REGION Network 19: TURUNKAN PRESSURE V 5
   RUNG wire#powerrail
      Contact( "DB106".Out_Step_17 )
      wire#w1
      I_Contact( "DB106".En_Step_19 )
      I_Contact( "Emergency" )
      Coil( "DB106".En_Step_18 )
   END_RUNG
   RUNG wire#powerrail
      Contact( "DB106".En_Step_18 )
   END_RUNG wire#w1
   // the same network as SCL:
   "DB106".En_Step_18 := ("DB106".Out_Step_17 OR "DB106".En_Step_18) AND NOT "DB106".En_Step_19 AND NOT "Emergency";
END_REGION

REGION Network 20: VB 5 OFF
   RUNG wire#powerrail
      Contact( "DB106".Out_Step_18 )
      { S7_Templates := "SrcType := Int" } LT_Contact(in1 := "Pressure vessel 5", in2 := 3)
      wire#w1
      I_Contact( "DB106".En_Step_20 )
      I_Contact( "Emergency" )
      Coil( "DB106".En_Step_19 )
   END_RUNG
   RUNG wire#powerrail
      Contact( "DB106".En_Step_19 )
   END_RUNG wire#w1
   // the same network as SCL:
   "DB106".En_Step_19 := (("DB106".Out_Step_18 AND ("Pressure vessel 5" < 3)) OR "DB106".En_Step_19) AND NOT "DB106".En_Step_20 AND NOT "Emergency";
END_REGION

REGION Network 21: VP 86 ON VP OFF
   RUNG wire#powerrail
      Contact( "DB106".Out_Step_19 )
      S_ODT(T_NO := "Tag_88", TV := S5T#4S, R :=, BI =>, RET_VAL =>)
      wire#w1
      I_Contact( "DB106".En_Step_21 )
      I_Contact( "Emergency" )
      Coil( "DB106".En_Step_20 )
   END_RUNG
   RUNG wire#powerrail
      Contact( "DB106".En_Step_20 )
   END_RUNG wire#w1
   // the same network as SCL:
   #_s5time1 := S_ODT(T_NO := "Tag_88", S := "DB106".Out_Step_19, TV := S5T#4S, Q => #_w1);
   "DB106".En_Step_20 := (#_w1 OR "DB106".En_Step_20) AND NOT "DB106".En_Step_21 AND NOT "Emergency";
END_REGION

REGION Network 22: VP 86 OFF VP 87 ON
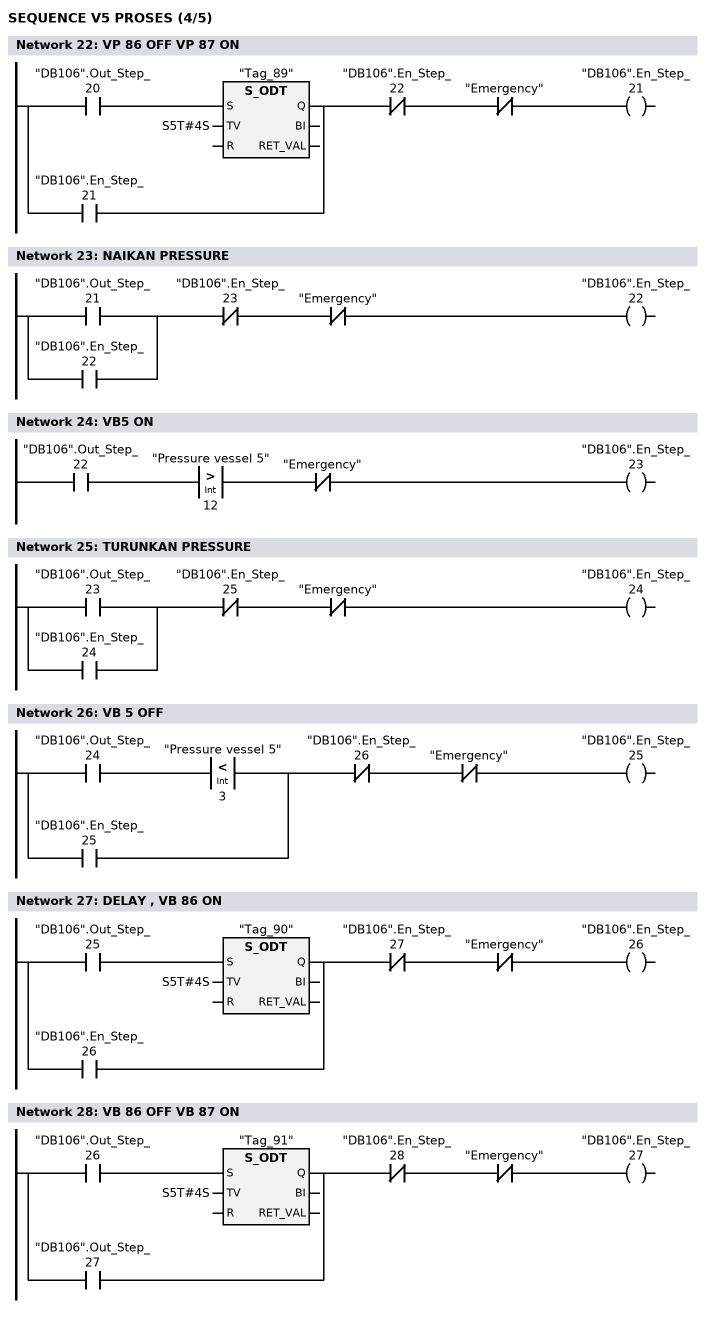
   RUNG wire#powerrail
      Contact( "DB106".Out_Step_20 )
      S_ODT(T_NO := "Tag_89", TV := S5T#4S, R :=, BI =>, RET_VAL =>)
      wire#w1
      I_Contact( "DB106".En_Step_22 )
      I_Contact( "Emergency" )
      Coil( "DB106".En_Step_21 )
   END_RUNG
   RUNG wire#powerrail
      Contact( "DB106".En_Step_21 )
   END_RUNG wire#w1
   // the same network as SCL:
   #_s5time1 := S_ODT(T_NO := "Tag_89", S := "DB106".Out_Step_20, TV := S5T#4S, Q => #_w1);
   "DB106".En_Step_21 := (#_w1 OR "DB106".En_Step_21) AND NOT "DB106".En_Step_22 AND NOT "Emergency";
END_REGION

REGION Network 23: NAIKAN PRESSURE
   RUNG wire#powerrail
      Contact( "DB106".Out_Step_21 )
      wire#w1
      I_Contact( "DB106".En_Step_23 )
      I_Contact( "Emergency" )
      Coil( "DB106".En_Step_22 )
   END_RUNG
   RUNG wire#powerrail
      Contact( "DB106".En_Step_22 )
   END_RUNG wire#w1
   // the same network as SCL:
   "DB106".En_Step_22 := ("DB106".Out_Step_21 OR "DB106".En_Step_22) AND NOT "DB106".En_Step_23 AND NOT "Emergency";
END_REGION

REGION Network 24: VB5 ON
   RUNG wire#powerrail
      Contact( "DB106".Out_Step_22 )
      { S7_Templates := "SrcType := Int" } GT_Contact(in1 := "Pressure vessel 5", in2 := 12)
      I_Contact( "Emergency" )
      Coil( "DB106".En_Step_23 )
   END_RUNG
   // the same network as SCL:
   "DB106".En_Step_23 := "DB106".Out_Step_22 AND ("Pressure vessel 5" > 12) AND NOT "Emergency";
END_REGION

REGION Network 25: TURUNKAN PRESSURE
   RUNG wire#powerrail
      Contact( "DB106".Out_Step_23 )
      wire#w1
      I_Contact( "DB106".En_Step_25 )
      I_Contact( "Emergency" )
      Coil( "DB106".En_Step_24 )
   END_RUNG
   RUNG wire#powerrail
      Contact( "DB106".En_Step_24 )
   END_RUNG wire#w1
   // the same network as SCL:
   "DB106".En_Step_24 := ("DB106".Out_Step_23 OR "DB106".En_Step_24) AND NOT "DB106".En_Step_25 AND NOT "Emergency";
END_REGION

REGION Network 26: VB 5 OFF
   RUNG wire#powerrail
      Contact( "DB106".Out_Step_24 )
      { S7_Templates := "SrcType := Int" } LT_Contact(in1 := "Pressure vessel 5", in2 := 3)
      wire#w1
      I_Contact( "DB106".En_Step_26 )
      I_Contact( "Emergency" )
      Coil( "DB106".En_Step_25 )
   END_RUNG
   RUNG wire#powerrail
      Contact( "DB106".En_Step_25 )
   END_RUNG wire#w1
   // the same network as SCL:
   "DB106".En_Step_25 := (("DB106".Out_Step_24 AND ("Pressure vessel 5" < 3)) OR "DB106".En_Step_25) AND NOT "DB106".En_Step_26 AND NOT "Emergency";
END_REGION

REGION Network 27: DELAY , VB 86 ON
   RUNG wire#powerrail
      Contact( "DB106".Out_Step_25 )
      S_ODT(T_NO := "Tag_90", TV := S5T#4S, R :=, BI =>, RET_VAL =>)
      wire#w1
      I_Contact( "DB106".En_Step_27 )
      I_Contact( "Emergency" )
      Coil( "DB106".En_Step_26 )
   END_RUNG
   RUNG wire#powerrail
      Contact( "DB106".En_Step_26 )
   END_RUNG wire#w1
   // the same network as SCL:
   #_s5time1 := S_ODT(T_NO := "Tag_90", S := "DB106".Out_Step_25, TV := S5T#4S, Q => #_w1);
   "DB106".En_Step_26 := (#_w1 OR "DB106".En_Step_26) AND NOT "DB106".En_Step_27 AND NOT "Emergency";
END_REGION

REGION Network 28: VB 86 OFF VB 87 ON
   RUNG wire#powerrail
      Contact( "DB106".Out_Step_26 )
      S_ODT(T_NO := "Tag_91", TV := S5T#4S, R :=, BI =>, RET_VAL =>)
      wire#w1
      I_Contact( "DB106".En_Step_28 )
      I_Contact( "Emergency" )
      Coil( "DB106".En_Step_27 )
   END_RUNG
   RUNG wire#powerrail
      Contact( "DB106".Out_Step_27 )
   END_RUNG wire#w1
   // the same network as SCL:
   #_s5time1 := S_ODT(T_NO := "Tag_91", S := "DB106".Out_Step_26, TV := S5T#4S, Q => #_w1);
   "DB106".En_Step_27 := (#_w1 OR "DB106".Out_Step_27) AND NOT "DB106".En_Step_28 AND NOT "Emergency";
END_REGION

REGION Network 29
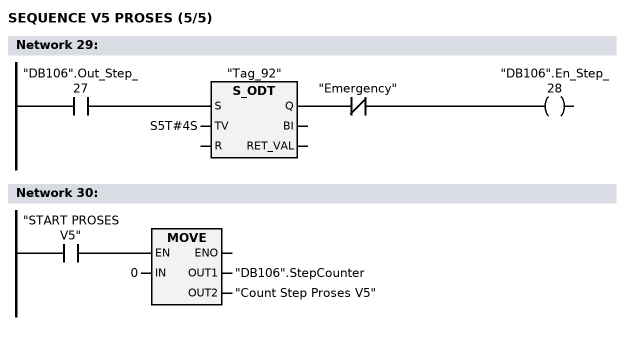
   RUNG wire#powerrail
      Contact( "DB106".Out_Step_27 )
      S_ODT(T_NO := "Tag_92", TV := S5T#4S, R :=, BI =>, RET_VAL =>)
      I_Contact( "Emergency" )
      Coil( "DB106".En_Step_28 )
   END_RUNG
   // the same network as SCL:
   #_s5time1 := S_ODT(T_NO := "Tag_92", S := "DB106".Out_Step_27, TV := S5T#4S, Q => #_w1);
   "DB106".En_Step_28 := #_w1 AND NOT "Emergency";
END_REGION

REGION Network 30
   RUNG wire#powerrail
      Contact( "START PROSES V5" )
      Move(in := 0, out1 => "DB106".StepCounter, out2 => "Count Step Proses V5")
   END_RUNG
   // the same network as SCL:
   IF "START PROSES V5" THEN
       "DB106".StepCounter := 0;
       "Count Step Proses V5" := 0;
   END_IF;
END_REGION
END_FUNCTION

FUNCTION "VESSEL 6 PROSES" : Void   // FC19, LAD
{ S7_Optimized_Access := 'TRUE' }
VERSION : 0.1
   VAR_TEMP   // added for the SCL form of the ladder/FBD networks
      _w1 : Bool;
      _w2 : Bool;
   END_VAR
BEGIN

REGION Network 1
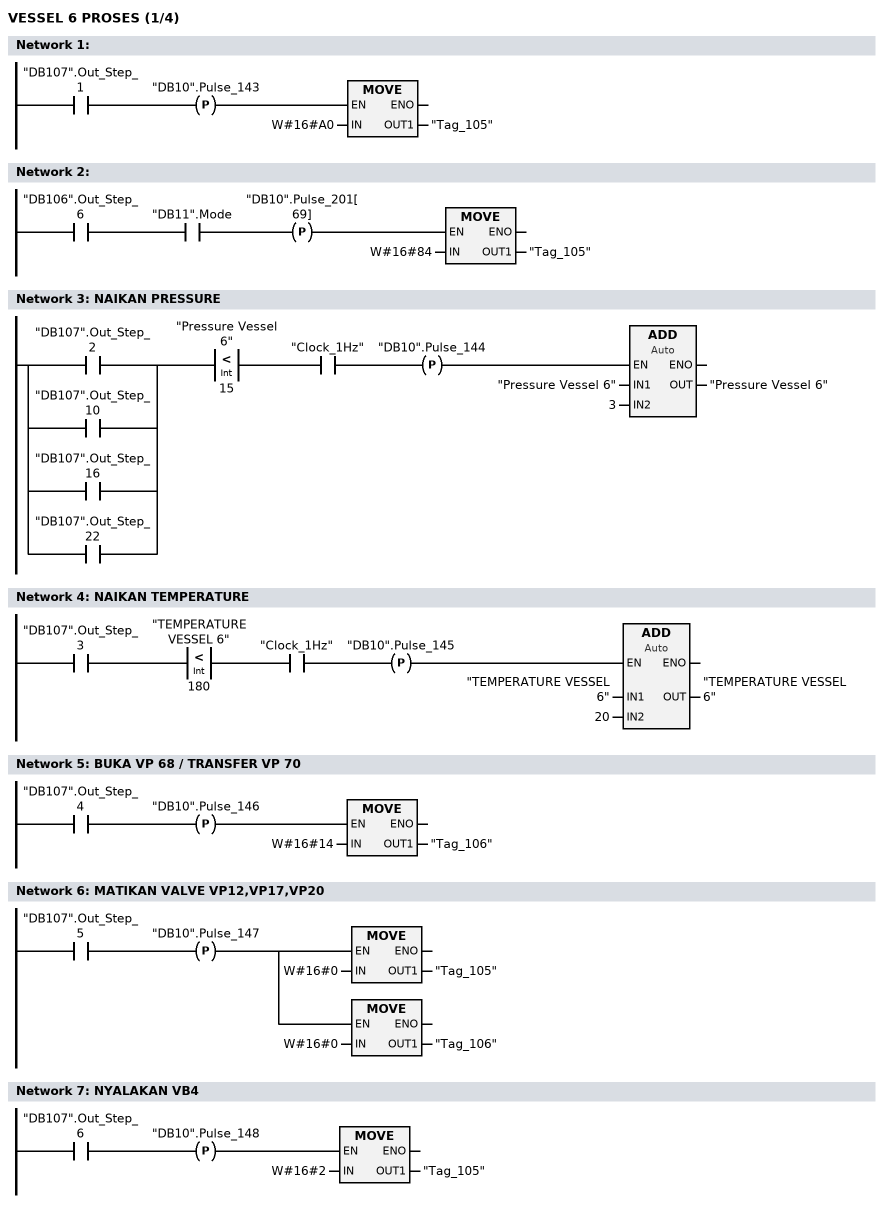
   RUNG wire#powerrail
      Contact( "DB107".Out_Step_1 )
      P_Trig( "DB10".Pulse_143 )
      Move(in := W#16#A0, out1 => "Tag_105")
   END_RUNG
   // the same network as SCL:
   #_w1 := "DB107".Out_Step_1 AND NOT "DB10".Pulse_143;   // rising edge
   "DB10".Pulse_143 := "DB107".Out_Step_1;
   IF #_w1 THEN "Tag_105" := W#16#A0; END_IF;
END_REGION

REGION Network 2
   RUNG wire#powerrail
      Contact( "DB106".Out_Step_6 )
      Contact( "DB11".Mode )
      P_Trig( "DB10".Pulse_201[69] )
      Move(in := W#16#84, out1 => "Tag_105")
   END_RUNG
   // the same network as SCL:
   #_w1 := "DB106".Out_Step_6 AND "DB11".Mode;
   #_w2 := #_w1 AND NOT "DB10".Pulse_201[69];   // rising edge
   "DB10".Pulse_201[69] := #_w1;
   IF #_w2 THEN "Tag_105" := W#16#84; END_IF;
END_REGION

REGION Network 3: NAIKAN PRESSURE
   RUNG wire#powerrail
      Contact( "DB107".Out_Step_2 )
      wire#w1
      { S7_Templates := "SrcType := Int" } LT_Contact(in1 := "Pressure Vessel 6", in2 := 15)
      Contact( "Clock_1Hz" )
      P_Trig( "DB10".Pulse_144 )
      Add(in1 := "Pressure Vessel 6", in2 := 3, out => "Pressure Vessel 6")
   END_RUNG
   RUNG wire#powerrail
      Contact( "DB107".Out_Step_10 )
   END_RUNG wire#w1
   RUNG wire#powerrail
      Contact( "DB107".Out_Step_16 )
   END_RUNG wire#w1
   RUNG wire#powerrail
      Contact( "DB107".Out_Step_22 )
   END_RUNG wire#w1
   // the same network as SCL:
   #_w1 := ("DB107".Out_Step_2 OR "DB107".Out_Step_10 OR "DB107".Out_Step_16 OR "DB107".Out_Step_22) AND ("Pressure Vessel 6" < 15) AND "Clock_1Hz";
   #_w2 := #_w1 AND NOT "DB10".Pulse_144;   // rising edge
   "DB10".Pulse_144 := #_w1;
   IF #_w2 THEN "Pressure Vessel 6" := "Pressure Vessel 6" + 3; END_IF;
END_REGION

REGION Network 4: NAIKAN TEMPERATURE
   RUNG wire#powerrail
      Contact( "DB107".Out_Step_3 )
      { S7_Templates := "SrcType := Int" } LT_Contact(in1 := "TEMPERATURE VESSEL 6", in2 := 180)
      Contact( "Clock_1Hz" )
      P_Trig( "DB10".Pulse_145 )
      Add(in1 := "TEMPERATURE VESSEL 6", in2 := 20, out => "TEMPERATURE VESSEL 6")
   END_RUNG
   // the same network as SCL:
   #_w1 := "DB107".Out_Step_3 AND ("TEMPERATURE VESSEL 6" < 180) AND "Clock_1Hz";
   #_w2 := #_w1 AND NOT "DB10".Pulse_145;   // rising edge
   "DB10".Pulse_145 := #_w1;
   IF #_w2 THEN "TEMPERATURE VESSEL 6" := "TEMPERATURE VESSEL 6" + 20; END_IF;
END_REGION

REGION Network 5: BUKA VP 68 / TRANSFER VP 70
   RUNG wire#powerrail
      Contact( "DB107".Out_Step_4 )
      P_Trig( "DB10".Pulse_146 )
      Move(in := W#16#14, out1 => "Tag_106")
   END_RUNG
   // the same network as SCL:
   #_w1 := "DB107".Out_Step_4 AND NOT "DB10".Pulse_146;   // rising edge
   "DB10".Pulse_146 := "DB107".Out_Step_4;
   IF #_w1 THEN "Tag_106" := W#16#14; END_IF;
END_REGION

REGION Network 6: MATIKAN VALVE VP12,VP17,VP20
   RUNG wire#powerrail
      Contact( "DB107".Out_Step_5 )
      P_Trig( "DB10".Pulse_147 )
      wire#w1
      Move(in := W#16#0, out1 => "Tag_105")
   END_RUNG
   RUNG wire#w1
      Move(in := W#16#0, out1 => "Tag_106")
   END_RUNG
   // the same network as SCL:
   #_w1 := "DB107".Out_Step_5 AND NOT "DB10".Pulse_147;   // rising edge
   "DB10".Pulse_147 := "DB107".Out_Step_5;
   IF #_w1 THEN
       "Tag_105" := W#16#0;
       "Tag_106" := W#16#0;
   END_IF;
END_REGION

REGION Network 7: NYALAKAN VB4
   RUNG wire#powerrail
      Contact( "DB107".Out_Step_6 )
      P_Trig( "DB10".Pulse_148 )
      Move(in := W#16#2, out1 => "Tag_105")
   END_RUNG
   // the same network as SCL:
   #_w1 := "DB107".Out_Step_6 AND NOT "DB10".Pulse_148;   // rising edge
   "DB10".Pulse_148 := "DB107".Out_Step_6;
   IF #_w1 THEN "Tag_105" := W#16#2; END_IF;
END_REGION

REGION Network 8: TURUNKAN PRESSURE
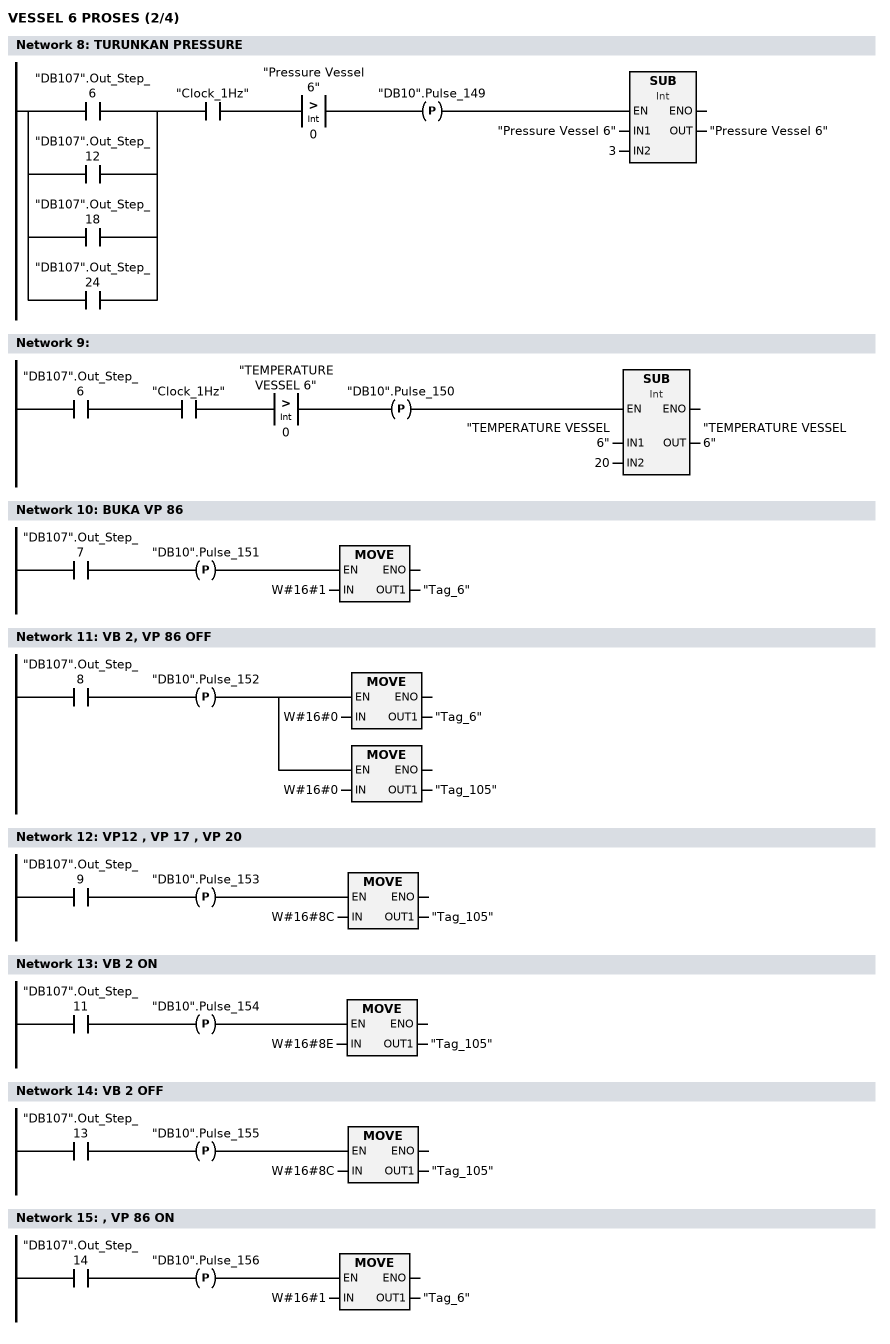
   RUNG wire#powerrail
      Contact( "DB107".Out_Step_6 )
      wire#w1
      Contact( "Clock_1Hz" )
      { S7_Templates := "SrcType := Int" } GT_Contact(in1 := "Pressure Vessel 6", in2 := 0)
      P_Trig( "DB10".Pulse_149 )
      { S7_Templates := "SrcType := Int" } Sub(in1 := "Pressure Vessel 6", in2 := 3, out => "Pressure Vessel 6")
   END_RUNG
   RUNG wire#powerrail
      Contact( "DB107".Out_Step_12 )
   END_RUNG wire#w1
   RUNG wire#powerrail
      Contact( "DB107".Out_Step_18 )
   END_RUNG wire#w1
   RUNG wire#powerrail
      Contact( "DB107".Out_Step_24 )
   END_RUNG wire#w1
   // the same network as SCL:
   #_w1 := ("DB107".Out_Step_6 OR "DB107".Out_Step_12 OR "DB107".Out_Step_18 OR "DB107".Out_Step_24) AND "Clock_1Hz" AND ("Pressure Vessel 6" > 0);
   #_w2 := #_w1 AND NOT "DB10".Pulse_149;   // rising edge
   "DB10".Pulse_149 := #_w1;
   IF #_w2 THEN "Pressure Vessel 6" := "Pressure Vessel 6" - 3; END_IF;
END_REGION

REGION Network 9
   RUNG wire#powerrail
      Contact( "DB107".Out_Step_6 )
      Contact( "Clock_1Hz" )
      { S7_Templates := "SrcType := Int" } GT_Contact(in1 := "TEMPERATURE VESSEL 6", in2 := 0)
      P_Trig( "DB10".Pulse_150 )
      { S7_Templates := "SrcType := Int" } Sub(in1 := "TEMPERATURE VESSEL 6", in2 := 20, out => "TEMPERATURE VESSEL 6")
   END_RUNG
   // the same network as SCL:
   #_w1 := "DB107".Out_Step_6 AND "Clock_1Hz" AND ("TEMPERATURE VESSEL 6" > 0);
   #_w2 := #_w1 AND NOT "DB10".Pulse_150;   // rising edge
   "DB10".Pulse_150 := #_w1;
   IF #_w2 THEN "TEMPERATURE VESSEL 6" := "TEMPERATURE VESSEL 6" - 20; END_IF;
END_REGION

REGION Network 10: BUKA VP 86
   RUNG wire#powerrail
      Contact( "DB107".Out_Step_7 )
      P_Trig( "DB10".Pulse_151 )
      Move(in := W#16#1, out1 => "Tag_6")
   END_RUNG
   // the same network as SCL:
   #_w1 := "DB107".Out_Step_7 AND NOT "DB10".Pulse_151;   // rising edge
   "DB10".Pulse_151 := "DB107".Out_Step_7;
   IF #_w1 THEN "Tag_6" := W#16#1; END_IF;
END_REGION

REGION Network 11: VB 2, VP 86 OFF
   RUNG wire#powerrail
      Contact( "DB107".Out_Step_8 )
      P_Trig( "DB10".Pulse_152 )
      wire#w1
      Move(in := W#16#0, out1 => "Tag_6")
   END_RUNG
   RUNG wire#w1
      Move(in := W#16#0, out1 => "Tag_105")
   END_RUNG
   // the same network as SCL:
   #_w1 := "DB107".Out_Step_8 AND NOT "DB10".Pulse_152;   // rising edge
   "DB10".Pulse_152 := "DB107".Out_Step_8;
   IF #_w1 THEN
       "Tag_6" := W#16#0;
       "Tag_105" := W#16#0;
   END_IF;
END_REGION

REGION Network 12: VP12 , VP 17 , VP 20
   RUNG wire#powerrail
      Contact( "DB107".Out_Step_9 )
      P_Trig( "DB10".Pulse_153 )
      Move(in := W#16#8C, out1 => "Tag_105")
   END_RUNG
   // the same network as SCL:
   #_w1 := "DB107".Out_Step_9 AND NOT "DB10".Pulse_153;   // rising edge
   "DB10".Pulse_153 := "DB107".Out_Step_9;
   IF #_w1 THEN "Tag_105" := W#16#8C; END_IF;
END_REGION

REGION Network 13: VB 2 ON
   RUNG wire#powerrail
      Contact( "DB107".Out_Step_11 )
      P_Trig( "DB10".Pulse_154 )
      Move(in := W#16#8E, out1 => "Tag_105")
   END_RUNG
   // the same network as SCL:
   #_w1 := "DB107".Out_Step_11 AND NOT "DB10".Pulse_154;   // rising edge
   "DB10".Pulse_154 := "DB107".Out_Step_11;
   IF #_w1 THEN "Tag_105" := W#16#8E; END_IF;
END_REGION

REGION Network 14: VB 2 OFF
   RUNG wire#powerrail
      Contact( "DB107".Out_Step_13 )
      P_Trig( "DB10".Pulse_155 )
      Move(in := W#16#8C, out1 => "Tag_105")
   END_RUNG
   // the same network as SCL:
   #_w1 := "DB107".Out_Step_13 AND NOT "DB10".Pulse_155;   // rising edge
   "DB10".Pulse_155 := "DB107".Out_Step_13;
   IF #_w1 THEN "Tag_105" := W#16#8C; END_IF;
END_REGION

REGION Network 15: , VP 86 ON
   RUNG wire#powerrail
      Contact( "DB107".Out_Step_14 )
      P_Trig( "DB10".Pulse_156 )
      Move(in := W#16#1, out1 => "Tag_6")
   END_RUNG
   // the same network as SCL:
   #_w1 := "DB107".Out_Step_14 AND NOT "DB10".Pulse_156;   // rising edge
   "DB10".Pulse_156 := "DB107".Out_Step_14;
   IF #_w1 THEN "Tag_6" := W#16#1; END_IF;
END_REGION

REGION Network 16: VP 86 OFF
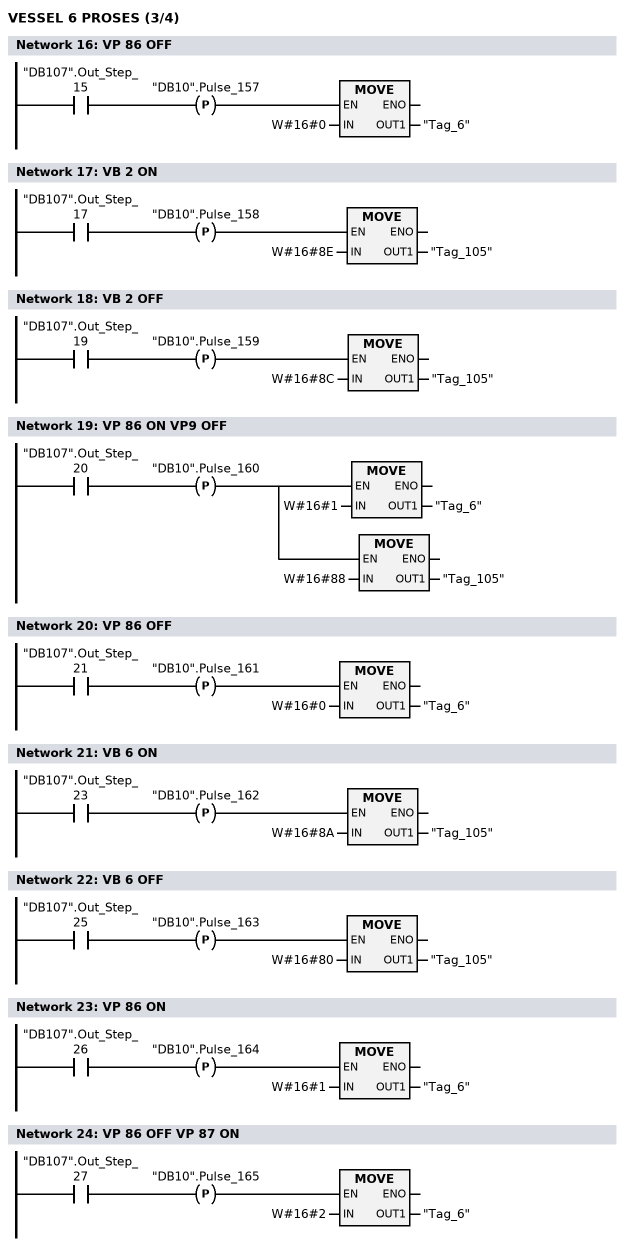
   RUNG wire#powerrail
      Contact( "DB107".Out_Step_15 )
      P_Trig( "DB10".Pulse_157 )
      Move(in := W#16#0, out1 => "Tag_6")
   END_RUNG
   // the same network as SCL:
   #_w1 := "DB107".Out_Step_15 AND NOT "DB10".Pulse_157;   // rising edge
   "DB10".Pulse_157 := "DB107".Out_Step_15;
   IF #_w1 THEN "Tag_6" := W#16#0; END_IF;
END_REGION

REGION Network 17: VB 2 ON
   RUNG wire#powerrail
      Contact( "DB107".Out_Step_17 )
      P_Trig( "DB10".Pulse_158 )
      Move(in := W#16#8E, out1 => "Tag_105")
   END_RUNG
   // the same network as SCL:
   #_w1 := "DB107".Out_Step_17 AND NOT "DB10".Pulse_158;   // rising edge
   "DB10".Pulse_158 := "DB107".Out_Step_17;
   IF #_w1 THEN "Tag_105" := W#16#8E; END_IF;
END_REGION

REGION Network 18: VB 2 OFF
   RUNG wire#powerrail
      Contact( "DB107".Out_Step_19 )
      P_Trig( "DB10".Pulse_159 )
      Move(in := W#16#8C, out1 => "Tag_105")
   END_RUNG
   // the same network as SCL:
   #_w1 := "DB107".Out_Step_19 AND NOT "DB10".Pulse_159;   // rising edge
   "DB10".Pulse_159 := "DB107".Out_Step_19;
   IF #_w1 THEN "Tag_105" := W#16#8C; END_IF;
END_REGION

REGION Network 19: VP 86 ON VP9 OFF
   RUNG wire#powerrail
      Contact( "DB107".Out_Step_20 )
      P_Trig( "DB10".Pulse_160 )
      wire#w1
      Move(in := W#16#1, out1 => "Tag_6")
   END_RUNG
   RUNG wire#w1
      Move(in := W#16#88, out1 => "Tag_105")
   END_RUNG
   // the same network as SCL:
   #_w1 := "DB107".Out_Step_20 AND NOT "DB10".Pulse_160;   // rising edge
   "DB10".Pulse_160 := "DB107".Out_Step_20;
   IF #_w1 THEN
       "Tag_6" := W#16#1;
       "Tag_105" := W#16#88;
   END_IF;
END_REGION

REGION Network 20: VP 86 OFF
   RUNG wire#powerrail
      Contact( "DB107".Out_Step_21 )
      P_Trig( "DB10".Pulse_161 )
      Move(in := W#16#0, out1 => "Tag_6")
   END_RUNG
   // the same network as SCL:
   #_w1 := "DB107".Out_Step_21 AND NOT "DB10".Pulse_161;   // rising edge
   "DB10".Pulse_161 := "DB107".Out_Step_21;
   IF #_w1 THEN "Tag_6" := W#16#0; END_IF;
END_REGION

REGION Network 21: VB 6 ON
   RUNG wire#powerrail
      Contact( "DB107".Out_Step_23 )
      P_Trig( "DB10".Pulse_162 )
      Move(in := W#16#8A, out1 => "Tag_105")
   END_RUNG
   // the same network as SCL:
   #_w1 := "DB107".Out_Step_23 AND NOT "DB10".Pulse_162;   // rising edge
   "DB10".Pulse_162 := "DB107".Out_Step_23;
   IF #_w1 THEN "Tag_105" := W#16#8A; END_IF;
END_REGION

REGION Network 22: VB 6 OFF
   RUNG wire#powerrail
      Contact( "DB107".Out_Step_25 )
      P_Trig( "DB10".Pulse_163 )
      Move(in := W#16#80, out1 => "Tag_105")
   END_RUNG
   // the same network as SCL:
   #_w1 := "DB107".Out_Step_25 AND NOT "DB10".Pulse_163;   // rising edge
   "DB10".Pulse_163 := "DB107".Out_Step_25;
   IF #_w1 THEN "Tag_105" := W#16#80; END_IF;
END_REGION

REGION Network 23: VP 86 ON
   RUNG wire#powerrail
      Contact( "DB107".Out_Step_26 )
      P_Trig( "DB10".Pulse_164 )
      Move(in := W#16#1, out1 => "Tag_6")
   END_RUNG
   // the same network as SCL:
   #_w1 := "DB107".Out_Step_26 AND NOT "DB10".Pulse_164;   // rising edge
   "DB10".Pulse_164 := "DB107".Out_Step_26;
   IF #_w1 THEN "Tag_6" := W#16#1; END_IF;
END_REGION

REGION Network 24: VP 86 OFF VP 87 ON
   RUNG wire#powerrail
      Contact( "DB107".Out_Step_27 )
      P_Trig( "DB10".Pulse_165 )
      Move(in := W#16#2, out1 => "Tag_6")
   END_RUNG
   // the same network as SCL:
   #_w1 := "DB107".Out_Step_27 AND NOT "DB10".Pulse_165;   // rising edge
   "DB10".Pulse_165 := "DB107".Out_Step_27;
   IF #_w1 THEN "Tag_6" := W#16#2; END_IF;
END_REGION

REGION Network 25: VP 87 OFF
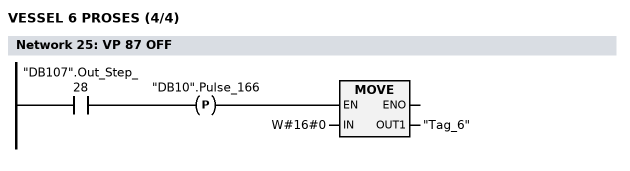
   RUNG wire#powerrail
      Contact( "DB107".Out_Step_28 )
      P_Trig( "DB10".Pulse_166 )
      Move(in := W#16#0, out1 => "Tag_6")
   END_RUNG
   // the same network as SCL:
   #_w1 := "DB107".Out_Step_28 AND NOT "DB10".Pulse_166;   // rising edge
   "DB10".Pulse_166 := "DB107".Out_Step_28;
   IF #_w1 THEN "Tag_6" := W#16#0; END_IF;
END_REGION
END_FUNCTION

FUNCTION "SEQUENCE V6 PROSES" : Void   // FC20, LAD
{ S7_Optimized_Access := 'TRUE' }
VERSION : 0.1
   VAR_TEMP   // added for the SCL form of the ladder/FBD networks
      _w1 : Bool;
      _w2 : Bool;
      _s5time1 : S5Time;
   END_VAR
BEGIN

REGION Network 1: START PROSES
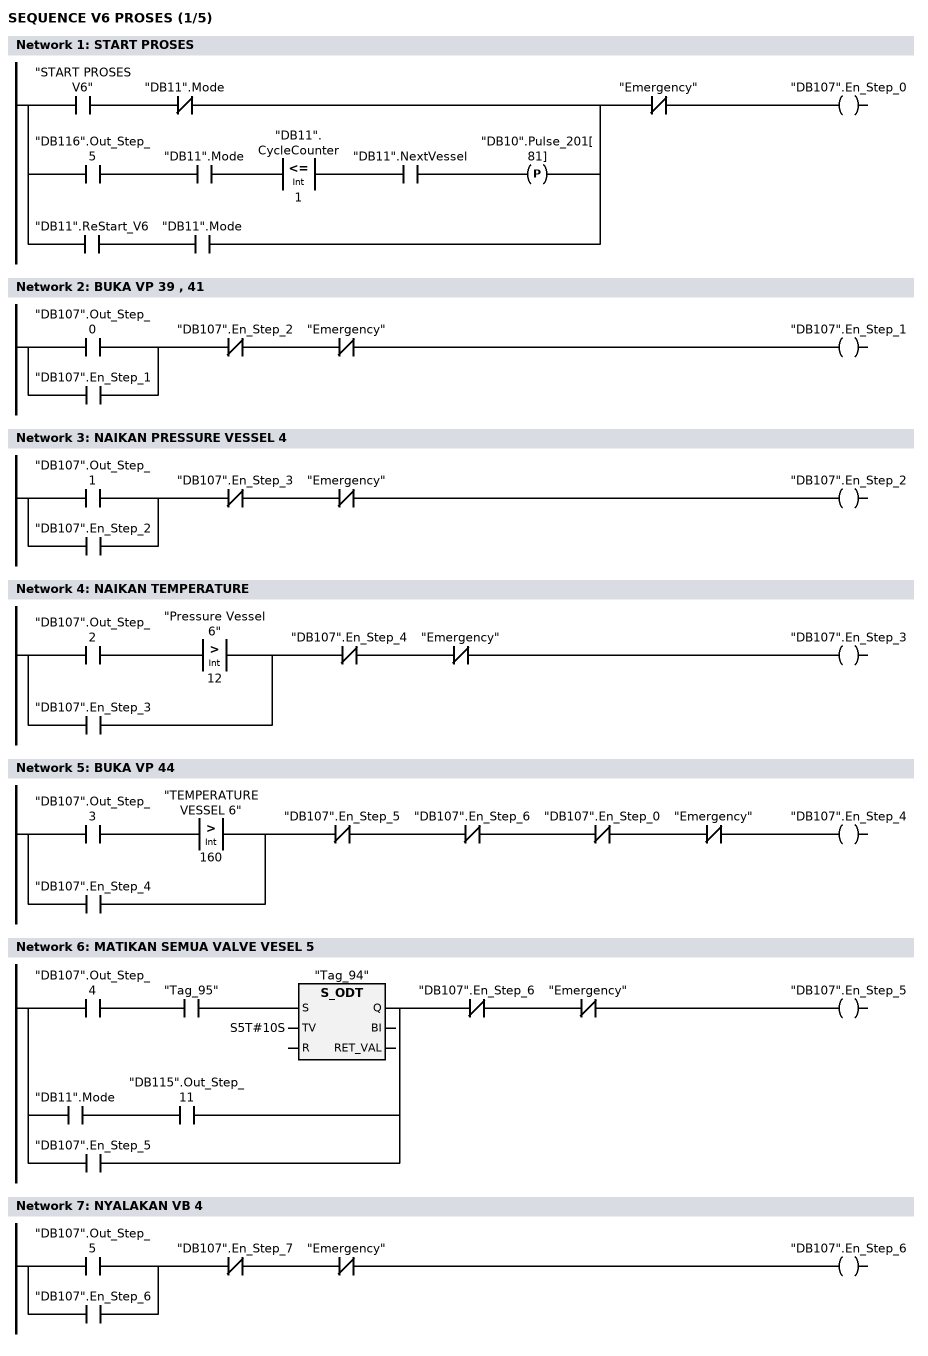
   RUNG wire#powerrail
      Contact( "START PROSES V6" )
      I_Contact( "DB11".Mode )
      wire#w1
      I_Contact( "Emergency" )
      Coil( "DB107".En_Step_0 )
   END_RUNG
   RUNG wire#powerrail
      Contact( "DB116".Out_Step_5 )
      Contact( "DB11".Mode )
      { S7_Templates := "SrcType := Int" } LE_Contact(in1 := "DB11".CycleCounter, in2 := 1)
      Contact( "DB11".NextVessel )
      P_Trig( "DB10".Pulse_201[81] )
   END_RUNG wire#w1
   RUNG wire#powerrail
      Contact( "DB11".ReStart_V6 )
      Contact( "DB11".Mode )
   END_RUNG wire#w1
   // the same network as SCL:
   #_w1 := "DB116".Out_Step_5 AND "DB11".Mode AND ("DB11".CycleCounter <= 1) AND "DB11".NextVessel;
   #_w2 := #_w1 AND NOT "DB10".Pulse_201[81];   // rising edge
   "DB10".Pulse_201[81] := #_w1;
   "DB107".En_Step_0 := (("START PROSES V6" AND NOT "DB11".Mode) OR #_w2 OR ("DB11".ReStart_V6 AND "DB11".Mode)) AND NOT "Emergency";
END_REGION

REGION Network 2: BUKA VP 39 , 41
   RUNG wire#powerrail
      Contact( "DB107".Out_Step_0 )
      wire#w1
      I_Contact( "DB107".En_Step_2 )
      I_Contact( "Emergency" )
      Coil( "DB107".En_Step_1 )
   END_RUNG
   RUNG wire#powerrail
      Contact( "DB107".En_Step_1 )
   END_RUNG wire#w1
   // the same network as SCL:
   "DB107".En_Step_1 := ("DB107".Out_Step_0 OR "DB107".En_Step_1) AND NOT "DB107".En_Step_2 AND NOT "Emergency";
END_REGION

REGION Network 3: NAIKAN PRESSURE VESSEL 4
   RUNG wire#powerrail
      Contact( "DB107".Out_Step_1 )
      wire#w1
      I_Contact( "DB107".En_Step_3 )
      I_Contact( "Emergency" )
      Coil( "DB107".En_Step_2 )
   END_RUNG
   RUNG wire#powerrail
      Contact( "DB107".En_Step_2 )
   END_RUNG wire#w1
   // the same network as SCL:
   "DB107".En_Step_2 := ("DB107".Out_Step_1 OR "DB107".En_Step_2) AND NOT "DB107".En_Step_3 AND NOT "Emergency";
END_REGION

REGION Network 4: NAIKAN TEMPERATURE
   RUNG wire#powerrail
      Contact( "DB107".Out_Step_2 )
      { S7_Templates := "SrcType := Int" } GT_Contact(in1 := "Pressure Vessel 6", in2 := 12)
      wire#w1
      I_Contact( "DB107".En_Step_4 )
      I_Contact( "Emergency" )
      Coil( "DB107".En_Step_3 )
   END_RUNG
   RUNG wire#powerrail
      Contact( "DB107".En_Step_3 )
   END_RUNG wire#w1
   // the same network as SCL:
   "DB107".En_Step_3 := (("DB107".Out_Step_2 AND ("Pressure Vessel 6" > 12)) OR "DB107".En_Step_3) AND NOT "DB107".En_Step_4 AND NOT "Emergency";
END_REGION

REGION Network 5: BUKA VP 44
   RUNG wire#powerrail
      Contact( "DB107".Out_Step_3 )
      { S7_Templates := "SrcType := Int" } GT_Contact(in1 := "TEMPERATURE VESSEL 6", in2 := 160)
      wire#w1
      I_Contact( "DB107".En_Step_5 )
      I_Contact( "DB107".En_Step_6 )
      I_Contact( "DB107".En_Step_0 )
      I_Contact( "Emergency" )
      Coil( "DB107".En_Step_4 )
   END_RUNG
   RUNG wire#powerrail
      Contact( "DB107".En_Step_4 )
   END_RUNG wire#w1
   // the same network as SCL:
   "DB107".En_Step_4 := (("DB107".Out_Step_3 AND ("TEMPERATURE VESSEL 6" > 160)) OR "DB107".En_Step_4) AND NOT "DB107".En_Step_5 AND NOT "DB107".En_Step_6 AND NOT "DB107".En_Step_0 AND NOT "Emergency";
END_REGION

REGION Network 6: MATIKAN SEMUA VALVE VESEL 5
   RUNG wire#powerrail
      Contact( "DB107".Out_Step_4 )
      Contact( "Tag_95" )
      S_ODT(T_NO := "Tag_94", TV := S5T#10S, R :=, BI =>, RET_VAL =>)
      wire#w1
      I_Contact( "DB107".En_Step_6 )
      I_Contact( "Emergency" )
      Coil( "DB107".En_Step_5 )
   END_RUNG
   RUNG wire#powerrail
      Contact( "DB11".Mode )
      Contact( "DB115".Out_Step_11 )
   END_RUNG wire#w1
   RUNG wire#powerrail
      Contact( "DB107".En_Step_5 )
   END_RUNG wire#w1
   // the same network as SCL:
   #_s5time1 := S_ODT(T_NO := "Tag_94", S := "DB107".Out_Step_4 AND "Tag_95", TV := S5T#10S, Q => #_w1);
   "DB107".En_Step_5 := (#_w1 OR ("DB11".Mode AND "DB115".Out_Step_11) OR "DB107".En_Step_5) AND NOT "DB107".En_Step_6 AND NOT "Emergency";
END_REGION

REGION Network 7: NYALAKAN VB 4
   RUNG wire#powerrail
      Contact( "DB107".Out_Step_5 )
      wire#w1
      I_Contact( "DB107".En_Step_7 )
      I_Contact( "Emergency" )
      Coil( "DB107".En_Step_6 )
   END_RUNG
   RUNG wire#powerrail
      Contact( "DB107".En_Step_6 )
   END_RUNG wire#w1
   // the same network as SCL:
   "DB107".En_Step_6 := ("DB107".Out_Step_5 OR "DB107".En_Step_6) AND NOT "DB107".En_Step_7 AND NOT "Emergency";
END_REGION

REGION Network 8
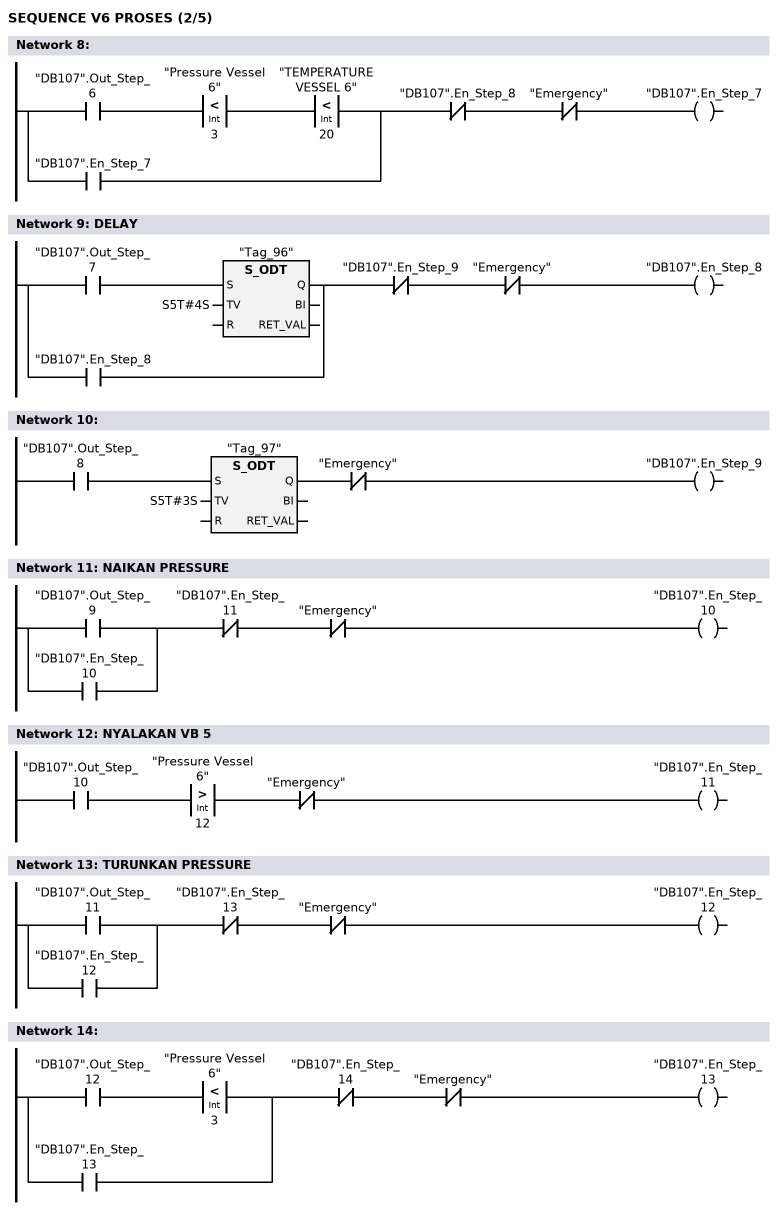
   RUNG wire#powerrail
      Contact( "DB107".Out_Step_6 )
      { S7_Templates := "SrcType := Int" } LT_Contact(in1 := "Pressure Vessel 6", in2 := 3)
      { S7_Templates := "SrcType := Int" } LT_Contact(in1 := "TEMPERATURE VESSEL 6", in2 := 20)
      wire#w1
      I_Contact( "DB107".En_Step_8 )
      I_Contact( "Emergency" )
      Coil( "DB107".En_Step_7 )
   END_RUNG
   RUNG wire#powerrail
      Contact( "DB107".En_Step_7 )
   END_RUNG wire#w1
   // the same network as SCL:
   "DB107".En_Step_7 := (("DB107".Out_Step_6 AND ("Pressure Vessel 6" < 3) AND ("TEMPERATURE VESSEL 6" < 20)) OR "DB107".En_Step_7) AND NOT "DB107".En_Step_8 AND NOT "Emergency";
END_REGION

REGION Network 9: DELAY
   RUNG wire#powerrail
      Contact( "DB107".Out_Step_7 )
      S_ODT(T_NO := "Tag_96", TV := S5T#4S, R :=, BI =>, RET_VAL =>)
      wire#w1
      I_Contact( "DB107".En_Step_9 )
      I_Contact( "Emergency" )
      Coil( "DB107".En_Step_8 )
   END_RUNG
   RUNG wire#powerrail
      Contact( "DB107".En_Step_8 )
   END_RUNG wire#w1
   // the same network as SCL:
   #_s5time1 := S_ODT(T_NO := "Tag_96", S := "DB107".Out_Step_7, TV := S5T#4S, Q => #_w1);
   "DB107".En_Step_8 := (#_w1 OR "DB107".En_Step_8) AND NOT "DB107".En_Step_9 AND NOT "Emergency";
END_REGION

REGION Network 10
   RUNG wire#powerrail
      Contact( "DB107".Out_Step_8 )
      S_ODT(T_NO := "Tag_97", TV := S5T#3S, R :=, BI =>, RET_VAL =>)
      I_Contact( "Emergency" )
      Coil( "DB107".En_Step_9 )
   END_RUNG
   // the same network as SCL:
   #_s5time1 := S_ODT(T_NO := "Tag_97", S := "DB107".Out_Step_8, TV := S5T#3S, Q => #_w1);
   "DB107".En_Step_9 := #_w1 AND NOT "Emergency";
END_REGION

REGION Network 11: NAIKAN PRESSURE
   RUNG wire#powerrail
      Contact( "DB107".Out_Step_9 )
      wire#w1
      I_Contact( "DB107".En_Step_11 )
      I_Contact( "Emergency" )
      Coil( "DB107".En_Step_10 )
   END_RUNG
   RUNG wire#powerrail
      Contact( "DB107".En_Step_10 )
   END_RUNG wire#w1
   // the same network as SCL:
   "DB107".En_Step_10 := ("DB107".Out_Step_9 OR "DB107".En_Step_10) AND NOT "DB107".En_Step_11 AND NOT "Emergency";
END_REGION

REGION Network 12: NYALAKAN VB 5
   RUNG wire#powerrail
      Contact( "DB107".Out_Step_10 )
      { S7_Templates := "SrcType := Int" } GT_Contact(in1 := "Pressure Vessel 6", in2 := 12)
      I_Contact( "Emergency" )
      Coil( "DB107".En_Step_11 )
   END_RUNG
   // the same network as SCL:
   "DB107".En_Step_11 := "DB107".Out_Step_10 AND ("Pressure Vessel 6" > 12) AND NOT "Emergency";
END_REGION

REGION Network 13: TURUNKAN PRESSURE
   RUNG wire#powerrail
      Contact( "DB107".Out_Step_11 )
      wire#w1
      I_Contact( "DB107".En_Step_13 )
      I_Contact( "Emergency" )
      Coil( "DB107".En_Step_12 )
   END_RUNG
   RUNG wire#powerrail
      Contact( "DB107".En_Step_12 )
   END_RUNG wire#w1
   // the same network as SCL:
   "DB107".En_Step_12 := ("DB107".Out_Step_11 OR "DB107".En_Step_12) AND NOT "DB107".En_Step_13 AND NOT "Emergency";
END_REGION

REGION Network 14
   RUNG wire#powerrail
      Contact( "DB107".Out_Step_12 )
      { S7_Templates := "SrcType := Int" } LT_Contact(in1 := "Pressure Vessel 6", in2 := 3)
      wire#w1
      I_Contact( "DB107".En_Step_14 )
      I_Contact( "Emergency" )
      Coil( "DB107".En_Step_13 )
   END_RUNG
   RUNG wire#powerrail
      Contact( "DB107".En_Step_13 )
   END_RUNG wire#w1
   // the same network as SCL:
   "DB107".En_Step_13 := (("DB107".Out_Step_12 AND ("Pressure Vessel 6" < 3)) OR "DB107".En_Step_13) AND NOT "DB107".En_Step_14 AND NOT "Emergency";
END_REGION

REGION Network 15
